   "Carrier_31_G120DControlWord.8" AT %I1911.0 : Bool;   // Bit_08_JOG_R
   "Carrier_31_G120DControlWord.9" AT %I1911.1 : Bool;   // Bit_09_JOG_L
   "Carrier_31_G120DControlWord.10" AT %I1911.2 : Bool;   // Bit_10_CONTR_PLC
   "Carrier_31_G120DControlWord.11" AT %I1911.3 : Bool;   // Bit_11_REVERSE
   "Carrier_31_G120DControlWord.12" AT %I1911.4 : Bool;   // Bit_12_BRAKE_RELEASE
   "Carrier_31_G120DControlWord.13" AT %I1911.5 : Bool;   // Bit_13_DDS
   "Carrier_31_G120DControlWord.14" AT %I1911.6 : Bool;   // Bit_14_DO0
   "Carrier_31_G120DControlWord.15" AT %I1911.7 : Bool;   // Bit_15_DO1
   "Carrier_31_G120DStatusWord" AT %IW1912 : Word;   // G120D_ZSW1_STATUS
   "Carrier_31_G120DStatusWord.0" AT %I1912.0 : Bool;   // Bit_00_READY_RUN
   "Carrier_31_G120DStatusWord.1" AT %I1912.1 : Bool;   // Bit_01_READY_ON
   "Carrier_31_G120DStatusWord.2" AT %I1912.2 : Bool;   // Bit_02_ENABLE
   "Carrier_31_G120DStatusWord.3" AT %I1912.3 : Bool;   // Bit_03_FAULT
   "Carrier_31_G120DStatusWord.4" AT %I1912.4 : Bool;   // Bit_04_OFF2
   "Carrier_31_G120DStatusWord.5" AT %I1912.5 : Bool;   // Bit_05_OFF3
   "Carrier_31_G120DStatusWord.6" AT %I1912.6 : Bool;   // Bit_06_LOCK_OUT
   "Carrier_31_G120DStatusWord.7" AT %I1912.7 : Bool;   // Bit_07_WARN
   "Carrier_31_G120DStatusWord.8" AT %I1913.0 : Bool;   // Bit_08_NO_DEVIATION
   "Carrier_31_G120DStatusWord.9" AT %I1913.1 : Bool;   // Bit_09_CONTR_PLC
   "Carrier_31_G120DStatusWord.10" AT %I1913.2 : Bool;   // Bit_10_F_MAX
   "Carrier_31_G120DStatusWord.11" AT %I1913.3 : Bool;   // Bit_11_LIMIT_REACHED
   "Carrier_31_G120DStatusWord.12" AT %I1913.4 : Bool;   // Bit_12_BRAKE_OPEN
   "Carrier_31_G120DStatusWord.13" AT %I1913.5 : Bool;   // Bit_13_NO_OVERTEMP
   "Carrier_31_G120DStatusWord.14" AT %I1913.6 : Bool;   // Bit_14_CW_CCW
   "Carrier_31_G120DStatusWord.15" AT %I1913.7 : Bool;   // Bit_15_OVERL
   "Carrier_31_Slot2_Input" AT %IW1914 : Word;   // SLOT 2 INPUT WORD
   "Carrier_31_CrashDetectSW" AT %I1914.0 : Bool;   // CRASH DETECT SW
   "Carrier_31_SpareSafetyInput(2_1)" AT %I1914.1 : Bool;   // SPARE SAFETY INPUT
   "Carrier_31_SpareSafetyInput(2_2)" AT %I1914.2 : Bool;   // SPARE SAFETY INPUT
   "Carrier_31_SpareSafetyInput(2_3)" AT %I1914.3 : Bool;   // SPARE SAFETY INPUT
   "Carrier_31_SpareSafetyInput(2_4)" AT %I1914.4 : Bool;   // SPARE SAFETY INPUT
   "Carrier_31_SpareSafetyInput(2_5)" AT %I1914.5 : Bool;   // SPARE SAFETY INPUT
   "Carrier_31_SpareSafetyInput(2_6)" AT %I1914.6 : Bool;   // SPARE SAFETY INPUT
   "Carrier_31_SpareSafetyInput(2_7)" AT %I1914.7 : Bool;   // SPARE SAFETY INPUT
   "Carrier_31_Slot3_SafetyOutput" AT %IW1915 : Word;   // SLOT 3 SAFETY OUTPUT WORD
   "Carrier_31_Crash_Detect_OK" AT %I1915.0 : Bool;   // CARRIER CRASH DETECT
   "Carrier_31_SpareSafetyOutput(3_1)" AT %I1915.1 : Bool;   // SPARE SAFETY OUTPUT
   "Carrier_31_SpareSafetyOutput(3_2)" AT %I1915.2 : Bool;   // SPARE SAFETY OUTPUT
   "Carrier_31_SpareSafetyOutput(3_3)" AT %I1915.3 : Bool;   // SPARE SAFETY OUTPUT
   "Carrier_31_SpareSafetyOutput(3_4)" AT %I1915.4 : Bool;   // SPARE SAFETY OUTPUT
   "Carrier_31_SpareSafetyOutput(3_5)" AT %I1915.5 : Bool;   // SPARE SAFETY OUTPUT
   "Carrier_31_SpareSafetyOutput(3_6)" AT %I1915.6 : Bool;   // SPARE SAFETY OUTPUT
   "Carrier_31_SpareSafetyOutput(3_7)" AT %I1915.7 : Bool;   // SPARE SAFETY OUTPUT
   "Carrier_31_Slot4_Input" AT %IW1916 : Word;   // SLOT 4 INPUT WORD
   "Carrier_31_480VPowerOn_MDCB1" AT %I1916.0 : Bool;   // 480 VAC POWER ON MDCB 1
   "Carrier_31_SpareInput(4_1)" AT %I1916.1 : Bool;   // SPARE INPUT
   "Carrier_31_SpareInput(4_2)" AT %I1916.2 : Bool;   // SPARE INPUT
   "Carrier_31_SitopSelectStatus" AT %I1916.3 : Bool;   // SITOP SELECT STATUS
   "Carrier_31_DCsupplyOnPSCB2" AT %I1916.4 : Bool;   // DC SUPPLY ON PSCB 2
   "Carrier_31_SpareInput(4_5)" AT %I1916.5 : Bool;   // SPARE INPUT
   "Carrier_31_SpareInput(4_6)" AT %I1916.6 : Bool;   // SPARE INPUT
   "Carrier_31_SpareInput(4_7)" AT %I1916.7 : Bool;   // SPARE INPUT
   "Carrier_31_PB1_ProdHoldLH" AT %I1917.0 : Bool;   // PB 1 PRODUCTION HOLD LH
   "Carrier_31_PB2_ResetLH" AT %I1917.1 : Bool;   // PB 2 RESET LH
   "Carrier_31_PB3_ProdHoldRH" AT %I1917.2 : Bool;   // PB 3 PRODUCTION HOLD RH
   "Carrier_31_PB4_ResetRH" AT %I1917.3 : Bool;   // PB 4 RESET RH
   "Carrier_31_SpareInput(4_14)" AT %I1917.4 : Bool;   // SPARE INPUT
   "Carrier_31_SpareInput(4_15)" AT %I1917.5 : Bool;   // SPARE INPUT
   "Carrier_31_SpareInput(4_16)" AT %I1917.6 : Bool;   // SPARE INPUT
   "Carrier_31_SpareInput(4_17)" AT %I1917.7 : Bool;   // SPARE INPUT
   "Carrier_31_Slot5_Output" AT %IW1918 : Word;   // SLOT 5 OUTPUT WORD
   "Carrier_31_IRD400_HMI_24VDC_ENABLE" AT %I1918.0 : Bool;   // IRD 400 PANEL HMI 24V DC POWER
   "Carrier_31_FaultLight_LH" AT %I1918.1 : Bool;   // FAULT LIGHT LH
   "Carrier_31_RunLight_LH" AT %I1918.2 : Bool;   // RUN LIGHT LH
   "Carrier_31_FaultLight_RH" AT %I1918.3 : Bool;   // FAULT LIGHT RH
   "Carrier_31_RunLight_RH" AT %I1918.4 : Bool;   // RUN LIGHT RH
   "Carrier_31_SpareOutput(5_5)" AT %I1918.5 : Bool;   // SPARE OUTPUT
   "Carrier_31_SpareOutput(5_6)" AT %I1918.6 : Bool;   // SPARE OUTPUT
   "Carrier_31_SpareOutput(5_7)" AT %I1918.7 : Bool;   // SPARE OUTPUT
   "Carrier_31_ActualSpeed" AT %IW1920 : Word;   // ACTUAL SPEED
   "Carrier_31_CarrierDriveAlarm" AT %IW1922 : Word;   // CARRIER DRIVE ALARM
   "Carrier_31_CarrierDriveWarning" AT %IW1924 : Word;   // CARRIER DRIVE WARNING
   "Carrier_32_Status" AT %IW1950 : Word;   // CARRIER STATUS WORD
   "Carrier_32_Status.0" AT %I1950.0 : Bool;   // HEARTBEAT
   "Carrier_32_Status.1" AT %I1950.1 : Bool;   // MANUAL
   "Carrier_32_Status.2" AT %I1950.2 : Bool;   // IN_AUTO
   "Carrier_32_Status.3" AT %I1950.3 : Bool;   // POSITIONING_COMPLETE
   "Carrier_32_Status.4" AT %I1950.4 : Bool;   // PRODUCTION HOLD
   "Carrier_32_Status.5" AT %I1950.5 : Bool;   // CARRIER MOVING FORWARD
   "Carrier_32_Status.6" AT %I1950.6 : Bool;   // CARRIER MOVING REVERSE
   "Carrier_32_Status.7" AT %I1950.7 : Bool;   // CARRIER FAULT
   "Carrier_32_Status.8" AT %I1951.0 : Bool;   // CRASH DETECT TRIPPED
   "Carrier_32_Status.9" AT %I1951.1 : Bool;
   "Carrier_32_Status.10" AT %I1951.2 : Bool;
   "Carrier_32_Status.11" AT %I1951.3 : Bool;
   "Carrier_32_Status.12" AT %I1951.4 : Bool;
   "Carrier_32_Status.13" AT %I1951.5 : Bool;
   "Carrier_32_Status.14" AT %I1951.6 : Bool;
   "Carrier_32_Status.15" AT %I1951.7 : Bool;
   "Carrier_32_SDCFaultCode" AT %IW1952 : Word;   // SDC FAULT CODE
   "Carrier_32_CarrierPosition" AT %ID1954 : DWord;   // CARRIER POSITION
   "Carrier_32_CarrierNumber" AT %IW1958 : Word;   // CARRIER NUMBER
   "Carrier_32_G120DControlWord" AT %IW1960 : Word;   // G120D_STW1_CONTROL
   "Carrier_32_G120DControlWord.0" AT %I1960.0 : Bool;   // Bit_00_ON
   "Carrier_32_G120DControlWord.1" AT %I1960.1 : Bool;   // Bit_01_AUS2_INH
   "Carrier_32_G120DControlWord.2" AT %I1960.2 : Bool;   // Bit_02_AUS3_STOP
   "Carrier_32_G120DControlWord.3" AT %I1960.3 : Bool;   // Bit_03_EN
   "Carrier_32_G120DControlWord.4" AT %I1960.4 : Bool;   // Bit_04_EN_RAMP
   "Carrier_32_G120DControlWord.5" AT %I1960.5 : Bool;   // Bit_05_START_RAMP
   "Carrier_32_G120DControlWord.6" AT %I1960.6 : Bool;   // Bit_06_SETPOINT
   "Carrier_32_G120DControlWord.7" AT %I1960.7 : Bool;   // Bit_07_RESET
   "Carrier_32_G120DControlWord.8" AT %I1961.0 : Bool;   // Bit_08_JOG_R
   "Carrier_32_G120DControlWord.9" AT %I1961.1 : Bool;   // Bit_09_JOG_L
   "Carrier_32_G120DControlWord.10" AT %I1961.2 : Bool;   // Bit_10_CONTR_PLC
   "Carrier_32_G120DControlWord.11" AT %I1961.3 : Bool;   // Bit_11_REVERSE
   "Carrier_32_G120DControlWord.12" AT %I1961.4 : Bool;   // Bit_12_BRAKE_RELEASE
   "Carrier_32_G120DControlWord.13" AT %I1961.5 : Bool;   // Bit_13_DDS
   "Carrier_32_G120DControlWord.14" AT %I1961.6 : Bool;   // Bit_14_DO0
   "Carrier_32_G120DControlWord.15" AT %I1961.7 : Bool;   // Bit_15_DO1
   "Carrier_32_G120DStatusWord" AT %IW1962 : Word;   // G120D_ZSW1_STATUS
   "Carrier_32_G120DStatusWord.0" AT %I1962.0 : Bool;   // Bit_00_READY_RUN
   "Carrier_32_G120DStatusWord.1" AT %I1962.1 : Bool;   // Bit_01_READY_ON
   "Carrier_32_G120DStatusWord.2" AT %I1962.2 : Bool;   // Bit_02_ENABLE
   "Carrier_32_G120DStatusWord.3" AT %I1962.3 : Bool;   // Bit_03_FAULT
   "Carrier_32_G120DStatusWord.4" AT %I1962.4 : Bool;   // Bit_04_OFF2
   "Carrier_32_G120DStatusWord.5" AT %I1962.5 : Bool;   // Bit_05_OFF3
   "Carrier_32_G120DStatusWord.6" AT %I1962.6 : Bool;   // Bit_06_LOCK_OUT
   "Carrier_32_G120DStatusWord.7" AT %I1962.7 : Bool;   // Bit_07_WARN
   "Carrier_32_G120DStatusWord.8" AT %I1963.0 : Bool;   // Bit_08_NO_DEVIATION
   "Carrier_32_G120DStatusWord.9" AT %I1963.1 : Bool;   // Bit_09_CONTR_PLC
   "Carrier_32_G120DStatusWord.10" AT %I1963.2 : Bool;   // Bit_10_F_MAX
   "Carrier_32_G120DStatusWord.11" AT %I1963.3 : Bool;   // Bit_11_LIMIT_REACHED
   "Carrier_32_G120DStatusWord.12" AT %I1963.4 : Bool;   // Bit_12_BRAKE_OPEN
   "Carrier_32_G120DStatusWord.13" AT %I1963.5 : Bool;   // Bit_13_NO_OVERTEMP
   "Carrier_32_G120DStatusWord.14" AT %I1963.6 : Bool;   // Bit_14_CW_CCW
   "Carrier_32_G120DStatusWord.15" AT %I1963.7 : Bool;   // Bit_15_OVERL
   "Carrier_32_Slot2_Input" AT %IW1964 : Word;   // SLOT 2 INPUT WORD
   "Carrier_32_CrashDetectSW" AT %I1964.0 : Bool;   // CRASH DETECT SW
   "Carrier_32_SpareSafetyInput(2_1)" AT %I1964.1 : Bool;   // SPARE SAFETY INPUT
   "Carrier_32_SpareSafetyInput(2_2)" AT %I1964.2 : Bool;   // SPARE SAFETY INPUT
   "Carrier_32_SpareSafetyInput(2_3)" AT %I1964.3 : Bool;   // SPARE SAFETY INPUT
   "Carrier_32_SpareSafetyInput(2_4)" AT %I1964.4 : Bool;   // SPARE SAFETY INPUT
   "Carrier_32_SpareSafetyInput(2_5)" AT %I1964.5 : Bool;   // SPARE SAFETY INPUT
   "Carrier_32_SpareSafetyInput(2_6)" AT %I1964.6 : Bool;   // SPARE SAFETY INPUT
   "Carrier_32_SpareSafetyInput(2_7)" AT %I1964.7 : Bool;   // SPARE SAFETY INPUT
   "Carrier_32_Slot3_SafetyOutput" AT %IW1965 : Word;   // SLOT 3 SAFETY OUTPUT WORD
   "Carrier_32_Crash_Detect_OK" AT %I1965.0 : Bool;   // CARRIER CRASH DETECT
   "Carrier_32_SpareSafetyOutput(3_1)" AT %I1965.1 : Bool;   // SPARE SAFETY OUTPUT
   "Carrier_32_SpareSafetyOutput(3_2)" AT %I1965.2 : Bool;   // SPARE SAFETY OUTPUT
   "Carrier_32_SpareSafetyOutput(3_3)" AT %I1965.3 : Bool;   // SPARE SAFETY OUTPUT
   "Carrier_32_SpareSafetyOutput(3_4)" AT %I1965.4 : Bool;   // SPARE SAFETY OUTPUT
   "Carrier_32_SpareSafetyOutput(3_5)" AT %I1965.5 : Bool;   // SPARE SAFETY OUTPUT
   "Carrier_32_SpareSafetyOutput(3_6)" AT %I1965.6 : Bool;   // SPARE SAFETY OUTPUT
   "Carrier_32_SpareSafetyOutput(3_7)" AT %I1965.7 : Bool;   // SPARE SAFETY OUTPUT
   "Carrier_32_Slot4_Input" AT %IW1966 : Word;   // SLOT 4 INPUT WORD
   "Carrier_32_480VPowerOn_MDCB1" AT %I1966.0 : Bool;   // 480 VAC POWER ON MDCB 1
   "Carrier_32_SpareInput(4_1)" AT %I1966.1 : Bool;   // SPARE INPUT
   "Carrier_32_SpareInput(4_2)" AT %I1966.2 : Bool;   // SPARE INPUT
   "Carrier_32_SitopSelectStatus" AT %I1966.3 : Bool;   // SITOP SELECT STATUS
   "Carrier_32_DCsupplyOnPSCB2" AT %I1966.4 : Bool;   // DC SUPPLY ON PSCB 2
   "Carrier_32_SpareInput(4_5)" AT %I1966.5 : Bool;   // SPARE INPUT
   "Carrier_32_SpareInput(4_6)" AT %I1966.6 : Bool;   // SPARE INPUT
   "Carrier_32_SpareInput(4_7)" AT %I1966.7 : Bool;   // SPARE INPUT
   "Carrier_32_PB1_ProdHoldLH" AT %I1967.0 : Bool;   // PB 1 PRODUCTION HOLD LH
   "Carrier_32_PB2_ResetLH" AT %I1967.1 : Bool;   // PB 2 RESET LH
   "Carrier_32_PB3_ProdHoldRH" AT %I1967.2 : Bool;   // PB 3 PRODUCTION HOLD RH
   "Carrier_32_PB4_ResetRH" AT %I1967.3 : Bool;   // PB 4 RESET RH
   "Carrier_32_SpareInput(4_14)" AT %I1967.4 : Bool;   // SPARE INPUT
   "Carrier_32_SpareInput(4_15)" AT %I1967.5 : Bool;   // SPARE INPUT
   "Carrier_32_SpareInput(4_16)" AT %I1967.6 : Bool;   // SPARE INPUT
   "Carrier_32_SpareInput(4_17)" AT %I1967.7 : Bool;   // SPARE INPUT
   "Carrier_32_Slot5_Output" AT %IW1968 : Word;   // SLOT 5 OUTPUT WORD
   "Carrier_32_IRD400_HMI_24VDC_ENABLE" AT %I1968.0 : Bool;   // IRD 400 PANEL HMI 24V DC POWER
   "Carrier_32_FaultLight_LH" AT %I1968.1 : Bool;   // FAULT LIGHT LH
   "Carrier_32_RunLight_LH" AT %I1968.2 : Bool;   // RUN LIGHT LH
   "Carrier_32_FaultLight_RH" AT %I1968.3 : Bool;   // FAULT LIGHT RH
   "Carrier_32_RunLight_RH" AT %I1968.4 : Bool;   // RUN LIGHT RH
   "Carrier_32_SpareOutput(5_5)" AT %I1968.5 : Bool;   // SPARE OUTPUT
   "Carrier_32_SpareOutput(5_6)" AT %I1968.6 : Bool;   // SPARE OUTPUT
   "Carrier_32_SpareOutput(5_7)" AT %I1968.7 : Bool;   // SPARE OUTPUT
   "Carrier_32_ActualSpeed" AT %IW1970 : Word;   // ACTUAL SPEED
   "Carrier_32_CarrierDriveAlarm" AT %IW1972 : Word;   // CARRIER DRIVE ALARM
   "Carrier_32_CarrierDriveWarning" AT %IW1974 : Word;   // CARRIER DRIVE WARNING
   "Carrier_33_Status" AT %IW2000 : Word;   // CARRIER STATUS WORD
   "Carrier_33_Status.0" AT %I2000.0 : Bool;   // HEARTBEAT
   "Carrier_33_Status.1" AT %I2000.1 : Bool;   // MANUAL
   "Carrier_33_Status.2" AT %I2000.2 : Bool;   // IN_AUTO
   "Carrier_33_Status.3" AT %I2000.3 : Bool;   // POSITIONING_COMPLETE
   "Carrier_33_Status.4" AT %I2000.4 : Bool;   // PRODUCTION HOLD
   "Carrier_33_Status.5" AT %I2000.5 : Bool;   // CARRIER MOVING FORWARD
   "Carrier_33_Status.6" AT %I2000.6 : Bool;   // CARRIER MOVING REVERSE
   "Carrier_33_Status.7" AT %I2000.7 : Bool;   // CARRIER FAULT
   "Carrier_33_Status.8" AT %I2001.0 : Bool;   // CRASH DETECT TRIPPED
   "Carrier_33_Status.9" AT %I2001.1 : Bool;
   "Carrier_33_Status.10" AT %I2001.2 : Bool;
   "Carrier_33_Status.11" AT %I2001.3 : Bool;
   "Carrier_33_Status.12" AT %I2001.4 : Bool;
   "Carrier_33_Status.13" AT %I2001.5 : Bool;
   "Carrier_33_Status.14" AT %I2001.6 : Bool;
   "Carrier_33_Status.15" AT %I2001.7 : Bool;
   "Carrier_33_SDCFaultCode" AT %IW2002 : Word;   // SDC FAULT CODE
   "Carrier_33_CarrierPosition" AT %ID2004 : DWord;   // CARRIER POSITION
   "Carrier_33_CarrierNumber" AT %IW2008 : Word;   // CARRIER NUMBER
   "Carrier_33_G120DControlWord" AT %IW2010 : Word;   // G120D_STW1_CONTROL
   "Carrier_33_G120DControlWord.0" AT %I2010.0 : Bool;   // Bit_00_ON
   "Carrier_33_G120DControlWord.1" AT %I2010.1 : Bool;   // Bit_01_AUS2_INH
   "Carrier_33_G120DControlWord.2" AT %I2010.2 : Bool;   // Bit_02_AUS3_STOP
   "Carrier_33_G120DControlWord.3" AT %I2010.3 : Bool;   // Bit_03_EN
   "Carrier_33_G120DControlWord.4" AT %I2010.4 : Bool;   // Bit_04_EN_RAMP
   "Carrier_33_G120DControlWord.5" AT %I2010.5 : Bool;   // Bit_05_START_RAMP
   "Carrier_33_G120DControlWord.6" AT %I2010.6 : Bool;   // Bit_06_SETPOINT
   "Carrier_33_G120DControlWord.7" AT %I2010.7 : Bool;   // Bit_07_RESET
   "Carrier_33_G120DControlWord.8" AT %I2011.0 : Bool;   // Bit_08_JOG_R
   "Carrier_33_G120DControlWord.9" AT %I2011.1 : Bool;   // Bit_09_JOG_L
   "Carrier_33_G120DControlWord.10" AT %I2011.2 : Bool;   // Bit_10_CONTR_PLC
   "Carrier_33_G120DControlWord.11" AT %I2011.3 : Bool;   // Bit_11_REVERSE
   "Carrier_33_G120DControlWord.12" AT %I2011.4 : Bool;   // Bit_12_BRAKE_RELEASE
   "Carrier_33_G120DControlWord.13" AT %I2011.5 : Bool;   // Bit_13_DDS
   "Carrier_33_G120DControlWord.14" AT %I2011.6 : Bool;   // Bit_14_DO0
   "Carrier_33_G120DControlWord.15" AT %I2011.7 : Bool;   // Bit_15_DO1
   "Carrier_33_G120DStatusWord" AT %IW2012 : Word;   // G120D_ZSW1_STATUS
   "Carrier_33_G120DStatusWord.0" AT %I2012.0 : Bool;   // Bit_00_READY_RUN
   "Carrier_33_G120DStatusWord.1" AT %I2012.1 : Bool;   // Bit_01_READY_ON
   "Carrier_33_G120DStatusWord.2" AT %I2012.2 : Bool;   // Bit_02_ENABLE
   "Carrier_33_G120DStatusWord.3" AT %I2012.3 : Bool;   // Bit_03_FAULT
   "Carrier_33_G120DStatusWord.4" AT %I2012.4 : Bool;   // Bit_04_OFF2
   "Carrier_33_G120DStatusWord.5" AT %I2012.5 : Bool;   // Bit_05_OFF3
   "Carrier_33_G120DStatusWord.6" AT %I2012.6 : Bool;   // Bit_06_LOCK_OUT
   "Carrier_33_G120DStatusWord.7" AT %I2012.7 : Bool;   // Bit_07_WARN
   "Carrier_33_G120DStatusWord.8" AT %I2013.0 : Bool;   // Bit_08_NO_DEVIATION
   "Carrier_33_G120DStatusWord.9" AT %I2013.1 : Bool;   // Bit_09_CONTR_PLC
   "Carrier_33_G120DStatusWord.10" AT %I2013.2 : Bool;   // Bit_10_F_MAX
   "Carrier_33_G120DStatusWord.11" AT %I2013.3 : Bool;   // Bit_11_LIMIT_REACHED
   "Carrier_33_G120DStatusWord.12" AT %I2013.4 : Bool;   // Bit_12_BRAKE_OPEN
   "Carrier_33_G120DStatusWord.13" AT %I2013.5 : Bool;   // Bit_13_NO_OVERTEMP
   "Carrier_33_G120DStatusWord.14" AT %I2013.6 : Bool;   // Bit_14_CW_CCW
   "Carrier_33_G120DStatusWord.15" AT %I2013.7 : Bool;   // Bit_15_OVERL
   "Carrier_33_Slot2_Input" AT %IW2014 : Word;   // SLOT 2 INPUT WORD
   "Carrier_33_CrashDetectSW" AT %I2014.0 : Bool;   // CRASH DETECT SW
   "Carrier_33_SpareSafetyInput(2_1)" AT %I2014.1 : Bool;   // SPARE SAFETY INPUT
   "Carrier_33_SpareSafetyInput(2_2)" AT %I2014.2 : Bool;   // SPARE SAFETY INPUT
   "Carrier_33_SpareSafetyInput(2_3)" AT %I2014.3 : Bool;   // SPARE SAFETY INPUT
   "Carrier_33_SpareSafetyInput(2_4)" AT %I2014.4 : Bool;   // SPARE SAFETY INPUT
   "Carrier_33_SpareSafetyInput(2_5)" AT %I2014.5 : Bool;   // SPARE SAFETY INPUT
   "Carrier_33_SpareSafetyInput(2_6)" AT %I2014.6 : Bool;   // SPARE SAFETY INPUT
   "Carrier_33_SpareSafetyInput(2_7)" AT %I2014.7 : Bool;   // SPARE SAFETY INPUT
   "Carrier_33_Slot3_SafetyOutput" AT %IW2015 : Word;   // SLOT 3 SAFETY OUTPUT WORD
   "Carrier_33_Crash_Detect_OK" AT %I2015.0 : Bool;   // CARRIER CRASH DETECT
   "Carrier_33_SpareSafetyOutput(3_1)" AT %I2015.1 : Bool;   // SPARE SAFETY OUTPUT
   "Carrier_33_SpareSafetyOutput(3_2)" AT %I2015.2 : Bool;   // SPARE SAFETY OUTPUT
   "Carrier_33_SpareSafetyOutput(3_3)" AT %I2015.3 : Bool;   // SPARE SAFETY OUTPUT
   "Carrier_33_SpareSafetyOutput(3_4)" AT %I2015.4 : Bool;   // SPARE SAFETY OUTPUT
   "Carrier_33_SpareSafetyOutput(3_5)" AT %I2015.5 : Bool;   // SPARE SAFETY OUTPUT
   "Carrier_33_SpareSafetyOutput(3_6)" AT %I2015.6 : Bool;   // SPARE SAFETY OUTPUT
   "Carrier_33_SpareSafetyOutput(3_7)" AT %I2015.7 : Bool;   // SPARE SAFETY OUTPUT
   "Carrier_33_Slot4_Input" AT %IW2016 : Word;   // SLOT 4 INPUT WORD
   "Carrier_33_480VPowerOn_MDCB1" AT %I2016.0 : Bool;   // 480 VAC POWER ON MDCB 1
   "Carrier_33_SpareInput(4_1)" AT %I2016.1 : Bool;   // SPARE INPUT
   "Carrier_33_SpareInput(4_2)" AT %I2016.2 : Bool;   // SPARE INPUT
   "Carrier_33_SitopSelectStatus" AT %I2016.3 : Bool;   // SITOP SELECT STATUS
   "Carrier_33_DCsupplyOnPSCB2" AT %I2016.4 : Bool;   // DC SUPPLY ON PSCB 2
   "Carrier_33_SpareInput(4_5)" AT %I2016.5 : Bool;   // SPARE INPUT
   "Carrier_33_SpareInput(4_6)" AT %I2016.6 : Bool;   // SPARE INPUT
   "Carrier_33_SpareInput(4_7)" AT %I2016.7 : Bool;   // SPARE INPUT
   "Carrier_33_PB1_ProdHoldLH" AT %I2017.0 : Bool;   // PB 1 PRODUCTION HOLD LH
   "Carrier_33_PB2_ResetLH" AT %I2017.1 : Bool;   // PB 2 RESET LH
   "Carrier_33_PB3_ProdHoldRH" AT %I2017.2 : Bool;   // PB 3 PRODUCTION HOLD RH
   "Carrier_33_PB4_ResetRH" AT %I2017.3 : Bool;   // PB 4 RESET RH
   "Carrier_33_SpareInput(4_14)" AT %I2017.4 : Bool;   // SPARE INPUT
   "Carrier_33_SpareInput(4_15)" AT %I2017.5 : Bool;   // SPARE INPUT
   "Carrier_33_SpareInput(4_16)" AT %I2017.6 : Bool;   // SPARE INPUT
   "Carrier_33_SpareInput(4_17)" AT %I2017.7 : Bool;   // SPARE INPUT
   "Carrier_33_Slot5_Output" AT %IW2018 : Word;   // SLOT 5 OUTPUT WORD
   "Carrier_33_IRD400_HMI_24VDC_ENABLE" AT %I2018.0 : Bool;   // IRD 400 PANEL HMI 24V DC POWER
   "Carrier_33_FaultLight_LH" AT %I2018.1 : Bool;   // FAULT LIGHT LH
   "Carrier_33_RunLight_LH" AT %I2018.2 : Bool;   // RUN LIGHT LH
   "Carrier_33_FaultLight_RH" AT %I2018.3 : Bool;   // FAULT LIGHT RH
   "Carrier_33_RunLight_RH" AT %I2018.4 : Bool;   // RUN LIGHT RH
   "Carrier_33_SpareOutput(5_5)" AT %I2018.5 : Bool;   // SPARE OUTPUT
   "Carrier_33_SpareOutput(5_6)" AT %I2018.6 : Bool;   // SPARE OUTPUT
   "Carrier_33_SpareOutput(5_7)" AT %I2018.7 : Bool;   // SPARE OUTPUT
   "Carrier_33_ActualSpeed" AT %IW2020 : Word;   // ACTUAL SPEED
   "Carrier_33_CarrierDriveAlarm" AT %IW2022 : Word;   // CARRIER DRIVE ALARM
   "Carrier_33_CarrierDriveWarning" AT %IW2024 : Word;   // CARRIER DRIVE WARNING
   "Carrier_34_Status" AT %IW2050 : Word;   // CARRIER STATUS WORD
   "Carrier_34_Status.0" AT %I2050.0 : Bool;   // HEARTBEAT
   "Carrier_34_Status.1" AT %I2050.1 : Bool;   // MANUAL
   "Carrier_34_Status.2" AT %I2050.2 : Bool;   // IN_AUTO
   "Carrier_34_Status.3" AT %I2050.3 : Bool;   // POSITIONING_COMPLETE
   "Carrier_34_Status.4" AT %I2050.4 : Bool;   // PRODUCTION HOLD
   "Carrier_34_Status.5" AT %I2050.5 : Bool;   // CARRIER MOVING FORWARD
   "Carrier_34_Status.6" AT %I2050.6 : Bool;   // CARRIER MOVING REVERSE
   "Carrier_34_Status.7" AT %I2050.7 : Bool;   // CARRIER FAULT
   "Carrier_34_Status.8" AT %I2051.0 : Bool;   // CRASH DETECT TRIPPED
   "Carrier_34_Status.9" AT %I2051.1 : Bool;
   "Carrier_34_Status.10" AT %I2051.2 : Bool;
   "Carrier_34_Status.11" AT %I2051.3 : Bool;
   "Carrier_34_Status.12" AT %I2051.4 : Bool;
   "Carrier_34_Status.13" AT %I2051.5 : Bool;
   "Carrier_34_Status.14" AT %I2051.6 : Bool;
   "Carrier_34_Status.15" AT %I2051.7 : Bool;
   "Carrier_34_SDCFaultCode" AT %IW2052 : Word;   // SDC FAULT CODE
   "Carrier_34_CarrierPosition" AT %ID2054 : DWord;   // CARRIER POSITION
   "Carrier_34_CarrierNumber" AT %IW2058 : Word;   // CARRIER NUMBER
   "Carrier_34_G120DControlWord" AT %IW2060 : Word;   // G120D_STW1_CONTROL
   "Carrier_34_G120DControlWord.0" AT %I2060.0 : Bool;   // Bit_00_ON
   "Carrier_34_G120DControlWord.1" AT %I2060.1 : Bool;   // Bit_01_AUS2_INH
   "Carrier_34_G120DControlWord.2" AT %I2060.2 : Bool;   // Bit_02_AUS3_STOP
   "Carrier_34_G120DControlWord.3" AT %I2060.3 : Bool;   // Bit_03_EN
   "Carrier_34_G120DControlWord.4" AT %I2060.4 : Bool;   // Bit_04_EN_RAMP
   "Carrier_34_G120DControlWord.5" AT %I2060.5 : Bool;   // Bit_05_START_RAMP
   "Carrier_34_G120DControlWord.6" AT %I2060.6 : Bool;   // Bit_06_SETPOINT
   "Carrier_34_G120DControlWord.7" AT %I2060.7 : Bool;   // Bit_07_RESET
   "Carrier_34_G120DControlWord.8" AT %I2061.0 : Bool;   // Bit_08_JOG_R
   "Carrier_34_G120DControlWord.9" AT %I2061.1 : Bool;   // Bit_09_JOG_L
   "Carrier_34_G120DControlWord.10" AT %I2061.2 : Bool;   // Bit_10_CONTR_PLC
   "Carrier_34_G120DControlWord.11" AT %I2061.3 : Bool;   // Bit_11_REVERSE
   "Carrier_34_G120DControlWord.12" AT %I2061.4 : Bool;   // Bit_12_BRAKE_RELEASE
   "Carrier_34_G120DControlWord.13" AT %I2061.5 : Bool;   // Bit_13_DDS
   "Carrier_34_G120DControlWord.14" AT %I2061.6 : Bool;   // Bit_14_DO0
   "Carrier_34_G120DControlWord.15" AT %I2061.7 : Bool;   // Bit_15_DO1
   "Carrier_34_G120DStatusWord" AT %IW2062 : Word;   // G120D_ZSW1_STATUS
   "Carrier_34_G120DStatusWord.0" AT %I2062.0 : Bool;   // Bit_00_READY_RUN
   "Carrier_34_G120DStatusWord.1" AT %I2062.1 : Bool;   // Bit_01_READY_ON
   "Carrier_34_G120DStatusWord.2" AT %I2062.2 : Bool;   // Bit_02_ENABLE
   "Carrier_34_G120DStatusWord.3" AT %I2062.3 : Bool;   // Bit_03_FAULT
   "Carrier_34_G120DStatusWord.4" AT %I2062.4 : Bool;   // Bit_04_OFF2
   "Carrier_34_G120DStatusWord.5" AT %I2062.5 : Bool;   // Bit_05_OFF3
   "Carrier_34_G120DStatusWord.6" AT %I2062.6 : Bool;   // Bit_06_LOCK_OUT
   "Carrier_34_G120DStatusWord.7" AT %I2062.7 : Bool;   // Bit_07_WARN
   "Carrier_34_G120DStatusWord.8" AT %I2063.0 : Bool;   // Bit_08_NO_DEVIATION
   "Carrier_34_G120DStatusWord.9" AT %I2063.1 : Bool;   // Bit_09_CONTR_PLC
   "Carrier_34_G120DStatusWord.10" AT %I2063.2 : Bool;   // Bit_10_F_MAX
   "Carrier_34_G120DStatusWord.11" AT %I2063.3 : Bool;   // Bit_11_LIMIT_REACHED
   "Carrier_34_G120DStatusWord.12" AT %I2063.4 : Bool;   // Bit_12_BRAKE_OPEN
   "Carrier_34_G120DStatusWord.13" AT %I2063.5 : Bool;   // Bit_13_NO_OVERTEMP
   "Carrier_34_G120DStatusWord.14" AT %I2063.6 : Bool;   // Bit_14_CW_CCW
   "Carrier_34_G120DStatusWord.15" AT %I2063.7 : Bool;   // Bit_15_OVERL
   "Carrier_34_Slot2_Input" AT %IW2064 : Word;   // SLOT 2 INPUT WORD
   "Carrier_34_CrashDetectSW" AT %I2064.0 : Bool;   // CRASH DETECT SW
   "Carrier_34_SpareSafetyInput(2_1)" AT %I2064.1 : Bool;   // SPARE SAFETY INPUT
   "Carrier_34_SpareSafetyInput(2_2)" AT %I2064.2 : Bool;   // SPARE SAFETY INPUT
   "Carrier_34_SpareSafetyInput(2_3)" AT %I2064.3 : Bool;   // SPARE SAFETY INPUT
   "Carrier_34_SpareSafetyInput(2_4)" AT %I2064.4 : Bool;   // SPARE SAFETY INPUT
   "Carrier_34_SpareSafetyInput(2_5)" AT %I2064.5 : Bool;   // SPARE SAFETY INPUT
   "Carrier_34_SpareSafetyInput(2_6)" AT %I2064.6 : Bool;   // SPARE SAFETY INPUT
   "Carrier_34_SpareSafetyInput(2_7)" AT %I2064.7 : Bool;   // SPARE SAFETY INPUT
   "Carrier_34_Slot3_SafetyOutput" AT %IW2065 : Word;   // SLOT 3 SAFETY OUTPUT WORD
   "Carrier_34_Crash_Detect_OK" AT %I2065.0 : Bool;   // CARRIER CRASH DETECT
   "Carrier_34_SpareSafetyOutput(3_1)" AT %I2065.1 : Bool;   // SPARE SAFETY OUTPUT
   "Carrier_34_SpareSafetyOutput(3_2)" AT %I2065.2 : Bool;   // SPARE SAFETY OUTPUT
   "Carrier_34_SpareSafetyOutput(3_3)" AT %I2065.3 : Bool;   // SPARE SAFETY OUTPUT
   "Carrier_34_SpareSafetyOutput(3_4)" AT %I2065.4 : Bool;   // SPARE SAFETY OUTPUT
   "Carrier_34_SpareSafetyOutput(3_5)" AT %I2065.5 : Bool;   // SPARE SAFETY OUTPUT
   "Carrier_34_SpareSafetyOutput(3_6)" AT %I2065.6 : Bool;   // SPARE SAFETY OUTPUT
   "Carrier_34_SpareSafetyOutput(3_7)" AT %I2065.7 : Bool;   // SPARE SAFETY OUTPUT
   "Carrier_34_Slot4_Input" AT %IW2066 : Word;   // SLOT 4 INPUT WORD
   "Carrier_34_480VPowerOn_MDCB1" AT %I2066.0 : Bool;   // 480 VAC POWER ON MDCB 1
   "Carrier_34_SpareInput(4_1)" AT %I2066.1 : Bool;   // SPARE INPUT
   "Carrier_34_SpareInput(4_2)" AT %I2066.2 : Bool;   // SPARE INPUT
   "Carrier_34_SitopSelectStatus" AT %I2066.3 : Bool;   // SITOP SELECT STATUS
   "Carrier_34_DCsupplyOnPSCB2" AT %I2066.4 : Bool;   // DC SUPPLY ON PSCB 2
   "Carrier_34_SpareInput(4_5)" AT %I2066.5 : Bool;   // SPARE INPUT
   "Carrier_34_SpareInput(4_6)" AT %I2066.6 : Bool;   // SPARE INPUT
   "Carrier_34_SpareInput(4_7)" AT %I2066.7 : Bool;   // SPARE INPUT
   "Carrier_34_PB1_ProdHoldLH" AT %I2067.0 : Bool;   // PB 1 PRODUCTION HOLD LH
   "Carrier_34_PB2_ResetLH" AT %I2067.1 : Bool;   // PB 2 RESET LH
   "Carrier_34_PB3_ProdHoldRH" AT %I2067.2 : Bool;   // PB 3 PRODUCTION HOLD RH
   "Carrier_34_PB4_ResetRH" AT %I2067.3 : Bool;   // PB 4 RESET RH
   "Carrier_34_SpareInput(4_14)" AT %I2067.4 : Bool;   // SPARE INPUT
   "Carrier_34_SpareInput(4_15)" AT %I2067.5 : Bool;   // SPARE INPUT
   "Carrier_34_SpareInput(4_16)" AT %I2067.6 : Bool;   // SPARE INPUT
   "Carrier_34_SpareInput(4_17)" AT %I2067.7 : Bool;   // SPARE INPUT
   "Carrier_34_Slot5_Output" AT %IW2068 : Word;   // SLOT 5 OUTPUT WORD
   "Carrier_34_IRD400_HMI_24VDC_ENABLE" AT %I2068.0 : Bool;   // IRD 400 PANEL HMI 24V DC POWER
   "Carrier_34_FaultLight_LH" AT %I2068.1 : Bool;   // FAULT LIGHT LH
   "Carrier_34_RunLight_LH" AT %I2068.2 : Bool;   // RUN LIGHT LH
   "Carrier_34_FaultLight_RH" AT %I2068.3 : Bool;   // FAULT LIGHT RH
   "Carrier_34_RunLight_RH" AT %I2068.4 : Bool;   // RUN LIGHT RH
   "Carrier_34_SpareOutput(5_5)" AT %I2068.5 : Bool;   // SPARE OUTPUT
   "Carrier_34_SpareOutput(5_6)" AT %I2068.6 : Bool;   // SPARE OUTPUT
   "Carrier_34_SpareOutput(5_7)" AT %I2068.7 : Bool;   // SPARE OUTPUT
   "Carrier_34_ActualSpeed" AT %IW2070 : Word;   // ACTUAL SPEED
   "Carrier_34_CarrierDriveAlarm" AT %IW2072 : Word;   // CARRIER DRIVE ALARM
   "Carrier_34_CarrierDriveWarning" AT %IW2074 : Word;   // CARRIER DRIVE WARNING
   "Carrier_35_Status" AT %IW2100 : Word;   // CARRIER STATUS WORD
   "Carrier_35_Status.0" AT %I2100.0 : Bool;   // HEARTBEAT
   "Carrier_35_Status.1" AT %I2100.1 : Bool;   // MANUAL
   "Carrier_35_Status.2" AT %I2100.2 : Bool;   // IN_AUTO
   "Carrier_35_Status.3" AT %I2100.3 : Bool;   // POSITIONING_COMPLETE
   "Carrier_35_Status.4" AT %I2100.4 : Bool;   // PRODUCTION HOLD
   "Carrier_35_Status.5" AT %I2100.5 : Bool;   // CARRIER MOVING FORWARD
   "Carrier_35_Status.6" AT %I2100.6 : Bool;   // CARRIER MOVING REVERSE
   "Carrier_35_Status.7" AT %I2100.7 : Bool;   // CARRIER FAULT
   "Carrier_35_Status.8" AT %I2101.0 : Bool;   // CRASH DETECT TRIPPED
   "Carrier_35_Status.9" AT %I2101.1 : Bool;
   "Carrier_35_Status.10" AT %I2101.2 : Bool;
   "Carrier_35_Status.11" AT %I2101.3 : Bool;
   "Carrier_35_Status.12" AT %I2101.4 : Bool;
   "Carrier_35_Status.13" AT %I2101.5 : Bool;
   "Carrier_35_Status.14" AT %I2101.6 : Bool;
   "Carrier_35_Status.15" AT %I2101.7 : Bool;
   "Carrier_35_SDCFaultCode" AT %IW2102 : Word;   // SDC FAULT CODE
   "Carrier_35_CarrierPosition" AT %ID2104 : DWord;   // CARRIER POSITION
   "Carrier_35_CarrierNumber" AT %IW2108 : Word;   // CARRIER NUMBER
   "Carrier_35_G120DControlWord" AT %IW2110 : Word;   // G120D_STW1_CONTROL
   "Carrier_35_G120DControlWord.0" AT %I2110.0 : Bool;   // Bit_00_ON
   "Carrier_35_G120DControlWord.1" AT %I2110.1 : Bool;   // Bit_01_AUS2_INH
   "Carrier_35_G120DControlWord.2" AT %I2110.2 : Bool;   // Bit_02_AUS3_STOP
   "Carrier_35_G120DControlWord.3" AT %I2110.3 : Bool;   // Bit_03_EN
   "Carrier_35_G120DControlWord.4" AT %I2110.4 : Bool;   // Bit_04_EN_RAMP
   "Carrier_35_G120DControlWord.5" AT %I2110.5 : Bool;   // Bit_05_START_RAMP
   "Carrier_35_G120DControlWord.6" AT %I2110.6 : Bool;   // Bit_06_SETPOINT
   "Carrier_35_G120DControlWord.7" AT %I2110.7 : Bool;   // Bit_07_RESET
   "Carrier_35_G120DControlWord.8" AT %I2111.0 : Bool;   // Bit_08_JOG_R
   "Carrier_35_G120DControlWord.9" AT %I2111.1 : Bool;   // Bit_09_JOG_L
   "Carrier_35_G120DControlWord.10" AT %I2111.2 : Bool;   // Bit_10_CONTR_PLC
   "Carrier_35_G120DControlWord.11" AT %I2111.3 : Bool;   // Bit_11_REVERSE
   "Carrier_35_G120DControlWord.12" AT %I2111.4 : Bool;   // Bit_12_BRAKE_RELEASE
   "Carrier_35_G120DControlWord.13" AT %I2111.5 : Bool;   // Bit_13_DDS
   "Carrier_35_G120DControlWord.14" AT %I2111.6 : Bool;   // Bit_14_DO0
   "Carrier_35_G120DControlWord.15" AT %I2111.7 : Bool;   // Bit_15_DO1
   "Carrier_35_G120DStatusWord" AT %IW2112 : Word;   // G120D_ZSW1_STATUS
   "Carrier_35_G120DStatusWord.0" AT %I2112.0 : Bool;   // Bit_00_READY_RUN
   "Carrier_35_G120DStatusWord.1" AT %I2112.1 : Bool;   // Bit_01_READY_ON
   "Carrier_35_G120DStatusWord.2" AT %I2112.2 : Bool;   // Bit_02_ENABLE
   "Carrier_35_G120DStatusWord.3" AT %I2112.3 : Bool;   // Bit_03_FAULT
   "Carrier_35_G120DStatusWord.4" AT %I2112.4 : Bool;   // Bit_04_OFF2
   "Carrier_35_G120DStatusWord.5" AT %I2112.5 : Bool;   // Bit_05_OFF3
   "Carrier_35_G120DStatusWord.6" AT %I2112.6 : Bool;   // Bit_06_LOCK_OUT
   "Carrier_35_G120DStatusWord.7" AT %I2112.7 : Bool;   // Bit_07_WARN
   "Carrier_35_G120DStatusWord.8" AT %I2113.0 : Bool;   // Bit_08_NO_DEVIATION
   "Carrier_35_G120DStatusWord.9" AT %I2113.1 : Bool;   // Bit_09_CONTR_PLC
   "Carrier_35_G120DStatusWord.10" AT %I2113.2 : Bool;   // Bit_10_F_MAX
   "Carrier_35_G120DStatusWord.11" AT %I2113.3 : Bool;   // Bit_11_LIMIT_REACHED
   "Carrier_35_G120DStatusWord.12" AT %I2113.4 : Bool;   // Bit_12_BRAKE_OPEN
   "Carrier_35_G120DStatusWord.13" AT %I2113.5 : Bool;   // Bit_13_NO_OVERTEMP
   "Carrier_35_G120DStatusWord.14" AT %I2113.6 : Bool;   // Bit_14_CW_CCW
   "Carrier_35_G120DStatusWord.15" AT %I2113.7 : Bool;   // Bit_15_OVERL
   "Carrier_35_Slot2_Input" AT %IW2114 : Word;   // SLOT 2 INPUT WORD
   "Carrier_35_CrashDetectSW" AT %I2114.0 : Bool;   // CRASH DETECT SW
   "Carrier_35_SpareSafetyInput(2_1)" AT %I2114.1 : Bool;   // SPARE SAFETY INPUT
   "Carrier_35_SpareSafetyInput(2_2)" AT %I2114.2 : Bool;   // SPARE SAFETY INPUT
   "Carrier_35_SpareSafetyInput(2_3)" AT %I2114.3 : Bool;   // SPARE SAFETY INPUT
   "Carrier_35_SpareSafetyInput(2_4)" AT %I2114.4 : Bool;   // SPARE SAFETY INPUT
   "Carrier_35_SpareSafetyInput(2_5)" AT %I2114.5 : Bool;   // SPARE SAFETY INPUT
   "Carrier_35_SpareSafetyInput(2_6)" AT %I2114.6 : Bool;   // SPARE SAFETY INPUT
   "Carrier_35_SpareSafetyInput(2_7)" AT %I2114.7 : Bool;   // SPARE SAFETY INPUT
   "Carrier_35_Slot3_SafetyOutput" AT %IW2115 : Word;   // SLOT 3 SAFETY OUTPUT WORD
   "Carrier_35_Crash_Detect_OK" AT %I2115.0 : Bool;   // CARRIER CRASH DETECT
   "Carrier_35_SpareSafetyOutput(3_1)" AT %I2115.1 : Bool;   // SPARE SAFETY OUTPUT
   "Carrier_35_SpareSafetyOutput(3_2)" AT %I2115.2 : Bool;   // SPARE SAFETY OUTPUT
   "Carrier_35_SpareSafetyOutput(3_3)" AT %I2115.3 : Bool;   // SPARE SAFETY OUTPUT
   "Carrier_35_SpareSafetyOutput(3_4)" AT %I2115.4 : Bool;   // SPARE SAFETY OUTPUT
   "Carrier_35_SpareSafetyOutput(3_5)" AT %I2115.5 : Bool;   // SPARE SAFETY OUTPUT
   "Carrier_35_SpareSafetyOutput(3_6)" AT %I2115.6 : Bool;   // SPARE SAFETY OUTPUT
   "Carrier_35_SpareSafetyOutput(3_7)" AT %I2115.7 : Bool;   // SPARE SAFETY OUTPUT
   "Carrier_35_Slot4_Input" AT %IW2116 : Word;   // SLOT 4 INPUT WORD
   "Carrier_35_480VPowerOn_MDCB1" AT %I2116.0 : Bool;   // 480 VAC POWER ON MDCB 1
   "Carrier_35_SpareInput(4_1)" AT %I2116.1 : Bool;   // SPARE INPUT
   "Carrier_35_SpareInput(4_2)" AT %I2116.2 : Bool;   // SPARE INPUT
   "Carrier_35_SitopSelectStatus" AT %I2116.3 : Bool;   // SITOP SELECT STATUS
   "Carrier_35_DCsupplyOnPSCB2" AT %I2116.4 : Bool;   // DC SUPPLY ON PSCB 2
   "Carrier_35_SpareInput(4_5)" AT %I2116.5 : Bool;   // SPARE INPUT
   "Carrier_35_SpareInput(4_6)" AT %I2116.6 : Bool;   // SPARE INPUT
   "Carrier_35_SpareInput(4_7)" AT %I2116.7 : Bool;   // SPARE INPUT
   "Carrier_35_PB1_ProdHoldLH" AT %I2117.0 : Bool;   // PB 1 PRODUCTION HOLD LH
   "Carrier_35_PB2_ResetLH" AT %I2117.1 : Bool;   // PB 2 RESET LH